   "2062_Warning_Data_BTCS_WARNING_WORD_13" : Word = PLC "2062_Warning_Data".BTCS_WARNING_WORD_13 AT %DB2062.DBW364, 1 s
   "2062_Warning_Data_BTCS_WARNING_WORD_14" : Word = PLC "2062_Warning_Data".BTCS_WARNING_WORD_14 AT %DB2062.DBW366, 1 s
   "2062_Warning_Data_BTCS_WARNING_WORD_15" : Word = PLC "2062_Warning_Data".BTCS_WARNING_WORD_15 AT %DB2062.DBW368, 1 s
   "2062_Warning_Data_BTCS_WARNING_WORD_16" : Word = PLC "2062_Warning_Data".BTCS_WARNING_WORD_16 AT %DB2062.DBW370, 1 s
   "2062_Warning_Data_BTCS_WARNING_WORD_2" : Word = PLC "2062_Warning_Data".BTCS_WARNING_WORD_02 AT %DB2062.DBW2, 1 s
   "2062_Warning_Data_BTCS_WARNING_WORD_3" : Word = PLC "2062_Warning_Data".BTCS_WARNING_WORD_03 AT %DB2062.DBW4, 1 s
   "2062_Warning_Data_BTCS_WARNING_WORD_4" : Word = PLC "2062_Warning_Data".BTCS_WARNING_WORD_04 AT %DB2062.DBW6, 1 s
   "2062_Warning_Data_BTCS_WARNING_WORD_5" : Word = PLC "2062_Warning_Data".BTCS_WARNING_WORD_05 AT %DB2062.DBW8, 1 s
   "2062_Warning_Data_BTCS_WARNING_WORD_6" : Word = PLC "2062_Warning_Data".BTCS_WARNING_WORD_06 AT %DB2062.DBW10, 1 s
   "2062_Warning_Data_BTCS_WARNING_WORD_7" : Word = PLC "2062_Warning_Data".BTCS_WARNING_WORD_07 AT %DB2062.DBW12, 1 s
   "2062_Warning_Data_BTCS_WARNING_WORD_8" : Word = PLC "2062_Warning_Data".BTCS_WARNING_WORD_08 AT %DB2062.DBW14, 1 s
   "2062_Warning_Data_Water Level Override 1P" : Bool = PLC "2062_Warning_Data"."Water Level Override 1P" AT %DB2062.DBX360.1, 1 s
   "2062_Warning_Data_Water Level Override 1S" : Bool = PLC "2062_Warning_Data"."Water Level Override 1S" AT %DB2062.DBX360.2, 1 s
   "2062_Warning_Data_Water Level Override 2P" : Bool = PLC "2062_Warning_Data"."Water Level Override 2P" AT %DB2062.DBX360.3, 1 s
   "2062_Warning_Data_Water Level Override 2S" : Bool = PLC "2062_Warning_Data"."Water Level Override 2S" AT %DB2062.DBX360.4, 1 s
   "2062_Warning_Data_Water Level Override 3P" : Bool = PLC "2062_Warning_Data"."Water Level Override 3P" AT %DB2062.DBX360.5, 1 s
   "2062_Warning_Data_Water Level Override 3S" : Bool = PLC "2062_Warning_Data"."Water Level Override 3S" AT %DB2062.DBX360.6, 1 s
   "2062_Warning_Data_Water Level Override 4P" : Bool = PLC "2062_Warning_Data"."Water Level Override 4P" AT %DB2062.DBX360.7, 1 s
   "2062_Warning_Data_Water Level Override 4S" : Bool = PLC "2062_Warning_Data"."Water Level Override 4S" AT %DB2062.DBX361.0, 1 s
   "2062_Warning_Data_Water Level Override 5P" : Bool = PLC "2062_Warning_Data"."Water Level Override 5P" AT %DB2062.DBX361.1, 1 s
   "2062_Warning_Data_Water Level Override 5S" : Bool = PLC "2062_Warning_Data"."Water Level Override 5S" AT %DB2062.DBX361.2, 1 s
   "2062_Warning_Data_Water Level Override 6P" : Bool = PLC "2062_Warning_Data"."Water Level Override 6P" AT %DB2062.DBX361.3, 1 s
   "2062_Warning_Data_Water Level Override 6S" : Bool = PLC "2062_Warning_Data"."Water Level Override 6S" AT %DB2062.DBX361.4, 1 s
   "2062_Warning_Data_Water Level Override APT" : Bool = PLC "2062_Warning_Data"."Water Level Override APT" AT %DB2062.DBX361.5, 1 s
   "2062_Warning_Data_Water Level Override FPT" : Bool = PLC "2062_Warning_Data"."Water Level Override FPT" AT %DB2062.DBX360.0, 1 s
   "2068_Sys_Status_Data_SAL_CNF_CHK" : Bool = PLC "2068_Sys_Status_Data".SAL_CNF_CHK, 100 ms
   "2068_Sys_Status_Data_SAL_VALID" : Bool = PLC "2068_Sys_Status_Data".SAL_VALID, 1 s
   "2086_Times_Alarm Enable Delay" : Time = PLC "2086_Times"."Alarm Enable Delay", 1 s
   "2086_Times_AT_DEOX_CNF_TIME" : Time = PLC "2086_Times".AT_DEOX_CNF_TIME AT %DB1.DBW0, 1 s
   "2086_Times_AT_REOX_CNF_TIME" : Time = PLC "2086_Times".AT_REOX_CNF_TIME AT %DB1.DBW0, 1 s
   "2086_Times_CV421_1S_MAX_TRVL_TIME" : Time = PLC "2086_Times".CV421_1S_MAX_TRVL_TIME, 1 s
   "2086_Times_CV421_2S_MAX_TRVL_TIME" : Time = PLC "2086_Times".CV421_2S_MAX_TRVL_TIME, 1 s
   "2086_Times_CV421_3S_MAX_TRVL_TIME" : Time = PLC "2086_Times".CV421_3S_MAX_TRVL_TIME, 1 s
   "2086_Times_CV421_4S_MAX_TRVL_TIME" : Time = PLC "2086_Times".CV421_4S_MAX_TRVL_TIME, 1 s
   "2086_Times_CV421_5S_MAX_TRVL_TIME" : Time = PLC "2086_Times".CV421_5S_MAX_TRVL_TIME, 1 s
   "2086_Times_CV421_6S_MAX_TRVL_TIME" : Time = PLC "2086_Times".CV421_6S_MAX_TRVL_TIME, 1 s
   "2086_Times_CV422_1P_MAX_TRVL_TIME" : Time = PLC "2086_Times".CV422_1P_MAX_TRVL_TIME, 1 s
   "2086_Times_CV422_2P_MAX_TRVL_TIME" : Time = PLC "2086_Times".CV422_2P_MAX_TRVL_TIME, 1 s
   "2086_Times_CV422_3P_MAX_TRVL_TIME" : Time = PLC "2086_Times".CV422_3P_MAX_TRVL_TIME, 1 s
   "2086_Times_CV422_4P_MAX_TRVL_TIME" : Time = PLC "2086_Times".CV422_4P_MAX_TRVL_TIME, 1 s
   "2086_Times_CV422_5P_MAX_TRVL_TIME" : Time = PLC "2086_Times".CV422_5P_MAX_TRVL_TIME, 1 s
   "2086_Times_CV422_6P_MAX_TRVL_TIME" : Time = PLC "2086_Times".CV422_6P_MAX_TRVL_TIME, 1 s
   "2086_Times_CV422_APT_MAX_TRVL_TIME" : Time = PLC "2086_Times".CV422_APT_MAX_TRVL_TIME, 1 s
   "2086_Times_CV422_FPT_MAX_TRVL_TIME" : Time = PLC "2086_Times".CV422_FPT_MAX_TRVL_TIME, 1 s
   "2086_Times_DEOX_PRE_GTT_CLS_DLY" : Time = PLC "2086_Times".DEOX_PRE_GTT_CLS_DLY AT %DB1.DBW0, 1 s
   "2086_Times_DEOX_PRE_GTT_OPN_DLY" : Time = PLC "2086_Times".DEOX_PRE_GTT_OPN_DLY AT %DB1.DBW0, 1 s
   "2086_Times_FIT417STAR Alarm Delay" : Time = PLC "2086_Times"."FIT417STAR Alarm Delay", 1 s
   "2086_Times_FIT418PORT Alarm Delay" : Time = PLC "2086_Times"."FIT418PORT Alarm Delay", 1 s
   "2086_Times_FIT419STAR Alarm Delay" : Time = PLC "2086_Times"."FIT419STAR Alarm Delay", 1 s
   "2086_Times_FIT420PORT Alarm Delay" : Time = PLC "2086_Times"."FIT420PORT Alarm Delay", 1 s
   "2086_Times_LS425 Port Alarm Delay" : Time = PLC "2086_Times"."LS425 Port Alarm Delay", 1 s
   "2086_Times_LS425 Star Alarm Delay" : Time = PLC "2086_Times"."LS425 Star Alarm Delay", 1 s
   "2086_Times_PIT424PORT Alarm Delay" : Time = PLC "2086_Times"."PIT424 Alarm Delay", 1 s
   "2086_Times_PS436 Alarm Delay" : Time = PLC "2086_Times"."PS436 Alarm Delay", 1 s
   "2086_Times_PT415PORT Alarm Delay" : Time = PLC "2086_Times"."PT415 Alarm Delay", 1 s
   "2086_Times_REOX_PRE_GTT_CLS_DLY" : Time = PLC "2086_Times".REOX_PRE_GTT_CLS_DLY AT %DB1.DBW0, 1 s
   "2086_Times_REOX_PRE_GTT_OPN_DLY" : Time = PLC "2086_Times".REOX_PRE_GTT_OPN_DLY AT %DB1.DBW0, 1 s
   "2086_Times_Tank Alarm Debounce" : Time = PLC "2086_Times"."Tank Alarm Reset Time", 1 s
   "2086_Times_TT426PORT Alarm Delay" : Time = PLC "2086_Times"."TT426_PORT_Alarm Delay", 1 s
   "2086_Times_TT426STAR Alarm Delay" : Time = PLC "2086_Times"."TT426_STAR_Alarm Delay", 1 s
   "21_FLOW_PRESSURE_SETPOINT_FIT_419_PRESSURE_SETPOINT" : Real = PLC "21_FLOW_PRESSURE_SETPOINT".FIT_419_PRESSURE_SETPOINT, 1 s
   "21_FLOW_PRESSURE_SETPOINT_FIT_420_PRESSURE_SETPOINT" : Real = PLC "21_FLOW_PRESSURE_SETPOINT".FIT_420_PRESSURE_SETPOINT, 1 s
   "2100_AUTO_SEQ_DB_SEQ_RNG" : Bool = PLC "2100_AUTO_SEQ_DB".SEQ_RNG, 1 s
   "2100_BTCS_CNTRL_DB_BTCS_STATE" : Int = PLC "2110_BTCS_CNTRL_DB".BTCS_STATE, 1 s
   "2100_BTCS_CNTRL_DB_BTCS_STEP" : Int = PLC "2110_BTCS_CNTRL_DB".BTCS_STEP, 1 s
   "2100_BTCS_CNTRL_DB_DE_OX_HRS" : Int = PLC "2110_BTCS_CNTRL_DB".DE_OX_HRS, 1 s
   "2100_BTCS_CNTRL_DB_DE_OX_MINS" : Int = PLC "2110_BTCS_CNTRL_DB".DE_OX_MINS, 1 s
   "2100_BTCS_CNTRL_DB_DE_OX_SP_HRS" : Int = PLC "2110_BTCS_CNTRL_DB".DE_OX_SP_HRS, 1 s
   "2100_BTCS_CNTRL_DB_DE_OX_SP_MINS" : Int = PLC "2110_BTCS_CNTRL_DB".DE_OX_SP_MINS, 1 s
   "2100_BTCS_CNTRL_DB_DWELL_HRS" : Int = PLC "2110_BTCS_CNTRL_DB".DWELL_HRS, 1 s
   "2100_BTCS_CNTRL_DB_DWELL_MINS" : Int = PLC "2110_BTCS_CNTRL_DB".DWELL_MINS, 1 s
   "2100_BTCS_CNTRL_DB_POST_DWELL_HRS" : Int = PLC "2110_BTCS_CNTRL_DB".POST_DWELL_HRS, 1 s
   "2100_BTCS_CNTRL_DB_POST_DWELL_MINS" : Int = PLC "2110_BTCS_CNTRL_DB".POST_DWELL_MINS, 1 s
   "2100_BTCS_CNTRL_DB_PRE_DWELL_HRS" : Int = PLC "2110_BTCS_CNTRL_DB".PRE_DWELL_HRS, 1 s
   "2100_BTCS_CNTRL_DB_PRE_DWELL_MINS" : Int = PLC "2110_BTCS_CNTRL_DB".PRE_DWELL_MINS, 1 s
   "2100_BTCS_CNTRL_DB_RE_OX_HRS" : Int = PLC "2110_BTCS_CNTRL_DB".RE_OX_HRS, 1 s
   "2100_BTCS_CNTRL_DB_RE_OX_MINS" : Int = PLC "2110_BTCS_CNTRL_DB".RE_OX_MINS, 1 s
   "2100_BTCS_CNTRL_DB_RE_OX_SP_HRS" : Int = PLC "2110_BTCS_CNTRL_DB".RE_OX_SP_HRS, 1 s
   "2100_BTCS_CNTRL_DB_RE_OX_SP_MINS" : Int = PLC "2110_BTCS_CNTRL_DB".RE_OX_SP_MINS, 1 s
   "2100_BTCS_CNTRL_DB_RMNG_SEQ_HRS" : Int = PLC "2110_BTCS_CNTRL_DB".RMNG_SEQ_HRS, 1 s
   "2100_BTCS_CNTRL_DB_RMNG_SEQ_MINS" : Int = PLC "2110_BTCS_CNTRL_DB".RMNG_SEQ_MINS, 1 s
   "2100_BTCS_CNTRL_DB_START_SEQ" : Bool = PLC "2110_BTCS_CNTRL_DB".START_SEQ, 1 s
   "2100_BTCS_CNTRL_DB_STOP_SEQ" : Bool = PLC "2110_BTCS_CNTRL_DB".STOP_SEQ, 1 s
   "2100_BTCS_CNTRL_DB_TOT_SEQ_HRS" : Int = PLC "2110_BTCS_CNTRL_DB".TOT_SEQ_HRS, 1 s
   "2100_BTCS_CNTRL_DB_TOT_SEQ_MINS" : Int = PLC "2110_BTCS_CNTRL_DB".TOT_SEQ_MINS, 1 s
   "2102_TIME_CALCS_DB_60X boost" : Bool = PLC "2102_TIME_CALCS_DB"."60X boost", 1 s
   "2102_TIME_CALCS_DB_DE_OX_MINS_RMNG" : Int = PLC "2102_TIME_CALCS_DB".DE_OX_MINS_RMNG, 1 s
   "2102_TIME_CALCS_DB_DE_OX_SP_MINS_RMNG" : Int = PLC "2102_TIME_CALCS_DB".DE_OX_SP_MINS_RMNG, 1 s
   "2102_TIME_CALCS_DB_DE_OX_SP_TMR_DN" : Bool = PLC "2102_TIME_CALCS_DB".DE_OX_SP_TMR_DN, 1 s
   "2102_TIME_CALCS_DB_DE_OX_TMR_DN" : Bool = PLC "2102_TIME_CALCS_DB".DE_OX_TMR_DN, 1 s
   "2102_TIME_CALCS_DB_DWELL_MINS_RMNG" : Int = PLC "2102_TIME_CALCS_DB".DWELL_MINS_RMNG, 1 s
   "2102_TIME_CALCS_DB_DWELL_TMR_DN" : Bool = PLC "2102_TIME_CALCS_DB".DWELL_TMR_DN, 1 s
   "2102_TIME_CALCS_DB_PHASE_DIFFERECE_MNS_REMNG" : Int = PLC "2102_TIME_CALCS_DB".PHASE_DIFFERECE_MNS_REMNG_De-Ox, 1 s
   "2102_TIME_CALCS_DB_POST_DWELL_MINS_RMNG" : Int = PLC "2102_TIME_CALCS_DB".POST_DWELL_MINS_RMNG, 1 s
   "2102_TIME_CALCS_DB_POST_DWELL_TMR_DN" : Bool = PLC "2102_TIME_CALCS_DB".POST_DWELL_TMR_DN, 1 s
   "2102_TIME_CALCS_DB_PRE_DWELL_MINS_RMNG" : Int = PLC "2102_TIME_CALCS_DB".PRE_DWELL_MINS_RMNG, 1 s
   "2102_TIME_CALCS_DB_PRE_DWELL_TMR_DN" : Bool = PLC "2102_TIME_CALCS_DB".PRE_DWELL_TMR_DN, 1 s
   "2102_TIME_CALCS_DB_PRE-DWEL MINS REMNG" : Int = PLC "2102_TIME_CALCS_DB"."PRE-DWEL MINS REMNG", 1 s
   "2102_TIME_CALCS_DB_PRE-DWEL_Warning 1" : Bool = PLC "2102_TIME_CALCS_DB"."PRE-DWEL_Warning 1", 500 ms
      on ChangeValue: "TimeRemainingToTreatment"()
   "2102_TIME_CALCS_DB_PRE-DWEL_Warning 2" : Bool = PLC "2102_TIME_CALCS_DB"."PRE-DWEL_Warning 2", 500 ms
      on ChangeValue: "TreatmentRequired"()
   "2102_TIME_CALCS_DB_PRE-DWEL_Warning 3" : Bool = PLC "2102_TIME_CALCS_DB"."PRE-DWEL_Warning 3", 1 s
   "2102_TIME_CALCS_DB_PRE-DWEL_Warning Min 1" : Int = PLC "2102_TIME_CALCS_DB"."PRE-DWEL_Warning Min 1", 1 s
   "2102_TIME_CALCS_DB_PRE-DWEL_Warning Min 2" : Int = PLC "2102_TIME_CALCS_DB"."PRE-DWEL_Warning Min 2", 1 s
   "2102_TIME_CALCS_DB_PRE-DWEL_Warning Min 3" : Int = PLC "2102_TIME_CALCS_DB"."PRE-DWEL_Warning Min 3", 1 s
   "2102_TIME_CALCS_DB_PRE-DWEL_Warning Reset 1" : Bool = PLC "2102_TIME_CALCS_DB"."PRE-DWEL_Warning Reset 1", 1 s
   "2102_TIME_CALCS_DB_PRE-DWEL_Warning Reset 2" : Bool = PLC "2102_TIME_CALCS_DB"."PRE-DWEL_Warning Reset 2", 1 s
   "2102_TIME_CALCS_DB_PRE-DWEL_Warning Reset 3" : Bool = PLC "2102_TIME_CALCS_DB"."PRE-DWEL_Warning Reset 3", 1 s
   "2102_TIME_CALCS_DB_RE_OX_MINS_RMNG" : Int = PLC "2102_TIME_CALCS_DB".RE_OX_MINS_RMNG, 1 s
   "2102_TIME_CALCS_DB_RE_OX_SP_MINS_RMNG" : Int = PLC "2102_TIME_CALCS_DB".RE_OX_SP_MINS_RMNG, 1 s
   "2102_TIME_CALCS_DB_RE_OX_SP_TMR_DN" : Bool = PLC "2102_TIME_CALCS_DB".RE_OX_SP_TMR_DN, 1 s
   "2102_TIME_CALCS_DB_RE_OX_TMR_DN" : Bool = PLC "2102_TIME_CALCS_DB".RE_OX_TMR_DN, 1 s
   "2102_TIME_CALCS_DB_Time_To_Treatment" : Int = PLC "2102_TIME_CALCS_DB".Time_To_Treatment, 1 s
   "2102_TIME_CALCS_DB_TIMES_VALID" : Bool = PLC "2102_TIME_CALCS_DB".TIMES_VALID, 1 s
   "2102_TIME_CALCS_DB_TOT_SEQ_DAYS" : Real = PLC "2102_TIME_CALCS_DB".TOT_SEQ_DAYS, 1 s
   "2102_TIME_CALCS_DB_TOT_SEQ_HRS_RMNG" : Int = PLC "2102_TIME_CALCS_DB".TOT_SEQ_HRS_RMNG, 1 s
   "2102_TIME_CALCS_DB_TOT_SEQ_MINS_RMNG" : Int = PLC "2102_TIME_CALCS_DB".TOT_SEQ_MINS_RMNG, 1 s
   "2102_TIME_CALCS_DB_Voyage_TIME_days" : Int = PLC "2102_TIME_CALCS_DB".Voyage_TIME_days, 1 s
   "2102_TIME_CALCS_DB_Voyage_TIME_hours" : Int = PLC "2102_TIME_CALCS_DB".Voyage_TIME_hours, 1 s
   "2102_TIME_CALCS_DB_Voyage_TIME_remaining_h" : Int = PLC "2102_TIME_CALCS_DB".Voyage_TIME_remaining_h, 1 s
   "2102_TIME_CALCS_DB_Voyage_TIME_remaining_m" : Int = PLC "2102_TIME_CALCS_DB".Voyage_TIME_remaining_m, 1 s
   "2110_BTCS_CNTRL_DB_PORT_TANK_STS" : Bool = PLC "2110_BTCS_CNTRL_DB".PORT_TANK_STS, 1 s
   "2110_BTCS_CNTRL_DB_RESET_ALL" : Bool = PLC "2110_BTCS_CNTRL_DB".RESET_ALL, 1 s
   "2110_BTCS_CNTRL_DB_STBD_TANK_STS" : Bool = PLC "2110_BTCS_CNTRL_DB".STBD_TANK_STS, 1 s
   "2115_VOYAGE_TIME_DAYS_VOYAGE_DAYS" : Real = PLC "2115_VOYAGE_TIME_DAYS".VOYAGE_DAYS, 1 s
   "40_TANKS_OP_DATA_RIO_02_VENT_A_2P" : Bool = PLC "40_TANKS_OP_DATA".RIO_02_VENT_A_2P AT %DB1.DBW0, 1 s
   "40_TANKS_OP_DATA_RIO_02_VENT_A_2S" : Bool = PLC "40_TANKS_OP_DATA".RIO_02_VENT_B_2S AT %DB1.DBW0, 1 s
   "40_TANKS_OP_DATA_RIO_02_VENT_B_2P" : Bool = PLC "40_TANKS_OP_DATA".RIO_02_VENT_B_2P AT %DB1.DBW0, 1 s
   "40_TANKS_OP_DATA_RIO_02_VENT_B_2S" : Bool = PLC "40_TANKS_OP_DATA".RIO_02_VENT_B_2P AT %DB1.DBW0, 1 s
   "502_ALM_ANALOG_IDB PIT 416_HIGH LEVEL VALUE (H)" : Real = PLC "502_ALM_ANALOG_IDB PIT 416"."HIGH LEVEL VALUE (H)" AT %DB65.DBD30, 1 s
   "502_ALM_ANALOG_IDB PIT 416_LOW LEVEL VALUE (L)" : Real = PLC "502_ALM_ANALOG_IDB PIT 416"."LOW LEVEL VALUE (L)" AT %DB65.DBD26, 1 s
   "502_ALM_ANALOG_IDB PIT 416_VERY HIGH LEVEL VALUE (HH)" : Real = PLC "502_ALM_ANALOG_IDB PIT 416"."VERY HIGH LEVEL VALUE (HH)" AT %DB65.DBD34, 1 s
   "502_ALM_ANALOG_IDB PIT 416_VERY LOW LEVEL VALUE (LL)" : Real = PLC "502_ALM_ANALOG_IDB PIT 416"."VERY LOW LEVEL VALUE (LL)" AT %DB65.DBD22, 1 s
   "503_WARNING CHCK_DB_2063_Alarm Word 12" : Word = PLC "503_WARNING CHCK_DB_2063"."Alarm Word 12", 1 s
   "503_WARNING CHCK_DB_2063_Alarm Word 13" : Word = PLC "503_WARNING CHCK_DB_2063"."Alarm Word 13", 1 s
   "503_WARNING CHCK_DB_2063_Alarm Word 14" : Word = PLC "503_WARNING CHCK_DB_2063"."Alarm Word 14", 1 s
   "503_WARNING CHCK_DB_2063_Alarm Word 15" : Word = PLC "503_WARNING CHCK_DB_2063"."Alarm Word 15", 1 s
   "503_WARNING CHCK_DB_2063_Alarm Word 16" : Word = PLC "503_WARNING CHCK_DB_2063"."Alarm Word 16", 1 s
   "504_Tank Grouping_DB2020_Boost" : Bool = PLC "504_Tank Grouping_DB2020".Boost, 1 s
   "504_Tank Grouping_DB2020_Cycle Length_ET" : Time = PLC "504_Tank Grouping_DB2020"."Cycle Length".ET, 1 s
   "504_Tank Grouping_DB2020_Cycle Period_ET" : Time = PLC "504_Tank Grouping_DB2020"."Cycle Period".ET, 1 s
   "504_Tank Grouping_DB2020_Diff Time Remain" : DInt = PLC "504_Tank Grouping_DB2020"."Diff Time Remain", 1 s
   "504_Tank Grouping_DB2020_GROUP ACTIV 1" : Bool = PLC "504_Tank Grouping_DB2020"."GROUP ACTIV 1", 1 s
   "504_Tank Grouping_DB2020_GROUP ACTIV 2" : Bool = PLC "504_Tank Grouping_DB2020"."GROUP ACTIV 2", 1 s
   "504_Tank Grouping_DB2020_GROUP ACTIV 3" : Bool = PLC "504_Tank Grouping_DB2020"."GROUP ACTIV 3", 1 s
   "504_Tank Grouping_DB2020_GROUP ACTIV 4" : Bool = PLC "504_Tank Grouping_DB2020"."GROUP ACTIV 4", 1 s
   "504_Tank Grouping_DB2020_GROUP ACTIV 5" : Bool = PLC "504_Tank Grouping_DB2020"."GROUP ACTIV 5", 1 s
   "504_Tank Grouping_DB2020_GROUP ACTIV 6" : Bool = PLC "504_Tank Grouping_DB2020"."GROUP ACTIV 6", 1 s
   "504_Tank Grouping_DB2020_GROUP ACTIV 7" : Bool = PLC "504_Tank Grouping_DB2020"."GROUP ACTIV 7", 1 s
   "504_Tank Grouping_DB2020_GROUP ACTIVE INT 1" : Bool = PLC "504_Tank Grouping_DB2020"."GROUP ACTIVE INT 1", 1 s
   "504_Tank Grouping_DB2020_GROUP ACTIVE INT 2" : Bool = PLC "504_Tank Grouping_DB2020"."GROUP ACTIVE INT 2", 1 s
   "504_Tank Grouping_DB2020_GROUP ACTIVE INT 3" : Bool = PLC "504_Tank Grouping_DB2020"."GROUP ACTIVE INT 3", 1 s
   "504_Tank Grouping_DB2020_GROUP ACTIVE INT 4" : Bool = PLC "504_Tank Grouping_DB2020"."GROUP ACTIVE INT 4", 1 s
   "504_Tank Grouping_DB2020_GROUP ACTIVE INT 5" : Bool = PLC "504_Tank Grouping_DB2020"."GROUP ACTIVE INT 5", 1 s
   "504_Tank Grouping_DB2020_GROUP ACTIVE INT 6" : Bool = PLC "504_Tank Grouping_DB2020"."GROUP ACTIVE INT 6", 1 s
   "504_Tank Grouping_DB2020_GROUP ACTIVE INT 7" : Bool = PLC "504_Tank Grouping_DB2020"."GROUP ACTIVE INT 7", 1 s
   "504_Tank Grouping_DB2020_GROUP of TANK 1" : Int = PLC "504_Tank Grouping_DB2020"."GROUP of TANK 1", 1 s
   "504_Tank Grouping_DB2020_GROUP of TANK 10" : Int = PLC "504_Tank Grouping_DB2020"."GROUP of TANK 10", 1 s
   "504_Tank Grouping_DB2020_GROUP of TANK 11" : Int = PLC "504_Tank Grouping_DB2020"."GROUP of TANK 11", 1 s
   "504_Tank Grouping_DB2020_GROUP of TANK 12" : Int = PLC "504_Tank Grouping_DB2020"."GROUP of TANK 12", 1 s
   "504_Tank Grouping_DB2020_GROUP of TANK 13" : Int = PLC "504_Tank Grouping_DB2020"."GROUP of TANK 13", 1 s
   "504_Tank Grouping_DB2020_GROUP of TANK 14" : Int = PLC "504_Tank Grouping_DB2020"."GROUP of TANK 14", 1 s
   "504_Tank Grouping_DB2020_GROUP of TANK 2" : Int = PLC "504_Tank Grouping_DB2020"."GROUP of TANK 2", 1 s
   "504_Tank Grouping_DB2020_GROUP of TANK 3" : Int = PLC "504_Tank Grouping_DB2020"."GROUP of TANK 3", 1 s
   "504_Tank Grouping_DB2020_GROUP of TANK 4" : Int = PLC "504_Tank Grouping_DB2020"."GROUP of TANK 4", 1 s
   "504_Tank Grouping_DB2020_GROUP of TANK 5" : Int = PLC "504_Tank Grouping_DB2020"."GROUP of TANK 5", 1 s
   "504_Tank Grouping_DB2020_GROUP of TANK 6" : Int = PLC "504_Tank Grouping_DB2020"."GROUP of TANK 6", 1 s
   "504_Tank Grouping_DB2020_GROUP of TANK 7" : Int = PLC "504_Tank Grouping_DB2020"."GROUP of TANK 7", 1 s
   "504_Tank Grouping_DB2020_GROUP of TANK 8" : Int = PLC "504_Tank Grouping_DB2020"."GROUP of TANK 8", 1 s
   "504_Tank Grouping_DB2020_GROUP of TANK 9" : Int = PLC "504_Tank Grouping_DB2020"."GROUP of TANK 9", 1 s
   "504_Tank Grouping_DB2020_GROUP SET" : Int = PLC "504_Tank Grouping_DB2020"."GROUP SET", 1 s
   "504_Tank Grouping_DB2020_O2 De-Ox Setpoint" : Real = PLC "504_Tank Grouping_DB2020"."O2 De-Ox Setpoint", 1 s
   "504_Tank Grouping_DB2020_Offset Timer_ET" : Time = PLC "504_Tank Grouping_DB2020"."Offset Timer".ET, 1 s
   "504_Tank Grouping_DB2020_RUN" : Bool = PLC "504_Tank Grouping_DB2020".RUN, 1 s
   "504_Tank Grouping_DB2020_RUN TANK 1" : Bool = PLC "504_Tank Grouping_DB2020"."RUN TANK 1", 1 s
   "504_Tank Grouping_DB2020_RUN TANK 10" : Bool = PLC "504_Tank Grouping_DB2020"."RUN TANK 10", 1 s
   "504_Tank Grouping_DB2020_RUN TANK 11" : Bool = PLC "504_Tank Grouping_DB2020"."RUN TANK 11", 1 s
   "504_Tank Grouping_DB2020_RUN TANK 12" : Bool = PLC "504_Tank Grouping_DB2020"."RUN TANK 12", 1 s
   "504_Tank Grouping_DB2020_RUN TANK 13" : Bool = PLC "504_Tank Grouping_DB2020"."RUN TANK 13", 1 s
   "504_Tank Grouping_DB2020_RUN TANK 14" : Bool = PLC "504_Tank Grouping_DB2020"."RUN TANK 14", 1 s
   "504_Tank Grouping_DB2020_RUN TANK 2" : Bool = PLC "504_Tank Grouping_DB2020"."RUN TANK 2", 1 s
   "504_Tank Grouping_DB2020_RUN TANK 3" : Bool = PLC "504_Tank Grouping_DB2020"."RUN TANK 3", 1 s
   "504_Tank Grouping_DB2020_RUN TANK 4" : Bool = PLC "504_Tank Grouping_DB2020"."RUN TANK 4", 1 s
   "504_Tank Grouping_DB2020_RUN TANK 5" : Bool = PLC "504_Tank Grouping_DB2020"."RUN TANK 5", 1 s
   "504_Tank Grouping_DB2020_RUN TANK 6" : Bool = PLC "504_Tank Grouping_DB2020"."RUN TANK 6", 1 s
   "504_Tank Grouping_DB2020_RUN TANK 7" : Bool = PLC "504_Tank Grouping_DB2020"."RUN TANK 7", 1 s
   "504_Tank Grouping_DB2020_RUN TANK 8" : Bool = PLC "504_Tank Grouping_DB2020"."RUN TANK 8", 1 s
   "504_Tank Grouping_DB2020_RUN TANK 9" : Bool = PLC "504_Tank Grouping_DB2020"."RUN TANK 9", 1 s
   "504_Tank Grouping_DB2020_Sequence Time Min Offset" : Time = PLC "504_Tank Grouping_DB2020"."Sequence Time m Offset", 1 s
   "504_Tank Grouping_DB2020_Sequence Time Min Offset_Int" : Real = PLC "504_Tank Grouping_DB2020"."Sequence Time m Offset_real", 1 s
   "504_Tank Grouping_DB2020_SetGroup" : Bool = PLC "504_Tank Grouping_DB2020".SetGroup, 1 s
   "504_Tank Grouping_DB2020_SetGroupSR" : Bool = PLC "504_Tank Grouping_DB2020".SetGroupSR, 1 s
   "504_Tank Grouping_DB2020_Tank1 Min Time_ET" : Time = PLC "504_Tank Grouping_DB2020"."Tank1 Min Time".ET, 1 s
   "504_Tank Grouping_DB2020_Tank10 Min Time_ET" : Time = PLC "504_Tank Grouping_DB2020"."Tank10 Min Time".ET, 1 s
   "504_Tank Grouping_DB2020_Tank12 Min Time_ET" : Time = PLC "504_Tank Grouping_DB2020"."Tank12 Min Time".ET, 1 s
   "504_Tank Grouping_DB2020_Tank13 Min Time_ET" : Time = PLC "504_Tank Grouping_DB2020"."Tank13 Min Time".ET, 1 s
   "504_Tank Grouping_DB2020_Tank14 Min Time_ET" : Time = PLC "504_Tank Grouping_DB2020"."Tank14 Min Time".ET, 1 s
   "504_Tank Grouping_DB2020_Tank2 Min Time_ET" : Time = PLC "504_Tank Grouping_DB2020"."Tank2 Min Time".ET, 1 s
   "504_Tank Grouping_DB2020_Tank3 Min Time_ET" : Time = PLC "504_Tank Grouping_DB2020"."Tank3 Min Time".ET, 1 s
   "504_Tank Grouping_DB2020_Tank4 Min Time_ET" : Time = PLC "504_Tank Grouping_DB2020"."Tank4 Min Time".ET, 1 s
   "504_Tank Grouping_DB2020_Tank5 Min Time_ET" : Time = PLC "504_Tank Grouping_DB2020"."Tank5 Min Time".ET, 1 s
   "504_Tank Grouping_DB2020_Tank6 Min Time_ET" : Time = PLC "504_Tank Grouping_DB2020"."Tank6 Min Time".ET, 1 s
   "504_Tank Grouping_DB2020_Tank7 Min Time_ET" : Time = PLC "504_Tank Grouping_DB2020"."Tank7 Min Time".ET, 1 s
   "504_Tank Grouping_DB2020_Tank8 Min Time_ET" : Time = PLC "504_Tank Grouping_DB2020"."Tank8 Min Time".ET, 1 s
   "504_Tank Grouping_DB2020_Tank9 Min Time_ET" : Time = PLC "504_Tank Grouping_DB2020"."Tank9 Min Time".ET, 1 s
   "504_Tank Grouping_DB2020_Time Left Tank_Time Left Tank 1" : Real = PLC "504_Tank Grouping_DB2020"."Time Left Tank"."Time Left Tank 1", 1 s
   "504_Tank Grouping_DB2020_Time Left Tank_Time Left Tank 10" : Real = PLC "504_Tank Grouping_DB2020"."Time Left Tank"."Time Left Tank 10", 1 s
   "504_Tank Grouping_DB2020_Time Left Tank_Time Left Tank 11" : Real = PLC "504_Tank Grouping_DB2020"."Time Left Tank"."Time Left Tank 11", 1 s
   "504_Tank Grouping_DB2020_Time Left Tank_Time Left Tank 12" : Real = PLC "504_Tank Grouping_DB2020"."Time Left Tank"."Time Left Tank 12", 1 s
   "504_Tank Grouping_DB2020_Time Left Tank_Time Left Tank 13" : Real = PLC "504_Tank Grouping_DB2020"."Time Left Tank"."Time Left Tank 13", 1 s
   "504_Tank Grouping_DB2020_Time Left Tank_Time Left Tank 14" : Real = PLC "504_Tank Grouping_DB2020"."Time Left Tank"."Time Left Tank 14", 1 s
   "504_Tank Grouping_DB2020_Time Left Tank_Time Left Tank 2" : Real = PLC "504_Tank Grouping_DB2020"."Time Left Tank"."Time Left Tank 2", 1 s
   "504_Tank Grouping_DB2020_Time Left Tank_Time Left Tank 3" : Real = PLC "504_Tank Grouping_DB2020"."Time Left Tank"."Time Left Tank 3", 1 s
   "504_Tank Grouping_DB2020_Time Left Tank_Time Left Tank 4" : Real = PLC "504_Tank Grouping_DB2020"."Time Left Tank"."Time Left Tank 4", 1 s
   "504_Tank Grouping_DB2020_Time Left Tank_Time Left Tank 5" : Real = PLC "504_Tank Grouping_DB2020"."Time Left Tank"."Time Left Tank 5", 1 s
   "504_Tank Grouping_DB2020_Time Left Tank_Time Left Tank 6" : Real = PLC "504_Tank Grouping_DB2020"."Time Left Tank"."Time Left Tank 6", 1 s
   "504_Tank Grouping_DB2020_Time Left Tank_Time Left Tank 7" : Real = PLC "504_Tank Grouping_DB2020"."Time Left Tank"."Time Left Tank 7", 1 s
   "504_Tank Grouping_DB2020_Time Left Tank_Time Left Tank 8" : Real = PLC "504_Tank Grouping_DB2020"."Time Left Tank"."Time Left Tank 8", 1 s
   "504_Tank Grouping_DB2020_Time Left Tank_Time Left Tank 9" : Real = PLC "504_Tank Grouping_DB2020"."Time Left Tank"."Time Left Tank 9", 1 s
   "504_Tank Grouping_DB2020_Valve Cycle_Enable" : Bool = PLC "504_Tank Grouping_DB2020"."Valve Cycle".Enable, 1 s
   "504_Tank Grouping_DB2020_Valve Cycle_Length" : Time = PLC "504_Tank Grouping_DB2020"."Valve Cycle".Length, 1 s
   "504_Tank Grouping_DB2020_Valve Cycle_Period" : Time = PLC "504_Tank Grouping_DB2020"."Valve Cycle".Period, 1 s
   "51_SLAVE_STATUS_RUNNING" : Bool = PLC "51_SLAVE_STATUS".RUNNING AT %DB51.DBX4.2, 1 s
   "60_Alarm_Data_ALRM_PRSNT" : Bool = PLC "60_Alarm_Data".ALRM_PRSNT AT %DB60.DBX32.0, 1 s
      on ChangeValue: "ALARM_Present"()
   "60_Alarm_Data_BC_ALARM_WORD_01" : Word = PLC "60_Alarm_Data".BC_ALARM_WORD_01 AT %DB60.DBW0, 1 s
   "60_Alarm_Data_BC_ALARM_WORD_02" : Word = PLC "60_Alarm_Data".BC_ALARM_WORD_02 AT %DB60.DBW2, 1 s
   "60_Alarm_Data_BC_ALARM_WORD_03" : Word = PLC "60_Alarm_Data".BC_ALARM_WORD_03 AT %DB60.DBW4, 1 s
   "60_Alarm_Data_BC_ALARM_WORD_04" : Word = PLC "60_Alarm_Data".BC_ALARM_WORD_04 AT %DB60.DBW6, 1 s
   "60_Alarm_Data_GCU_ALARM_WORD_01" : Word = PLC "60_Alarm_Data".GCU_ALARM_WORD_01 AT %DB60.DBW0, 1 s
   "60_Alarm_Data_GCU_ALARM_WORD_02" : Word = PLC "60_Alarm_Data".GCU_ALARM_WORD_02 AT %DB60.DBW2, 1 s
   "60_Alarm_Data_GCU_ALARM_WORD_03" : Word = PLC "60_Alarm_Data".GCU_ALARM_WORD_03 AT %DB60.DBW4, 1 s
   "60_Alarm_Data_GCU_ALARM_WORD_04" : Word = PLC "60_Alarm_Data".GCU_ALARM_WORD_04 AT %DB60.DBW6, 1 s
   "60_Alarm_Data_GCU_ALARM_WORD_05" : Word = PLC "60_Alarm_Data".GCU_ALARM_WORD_05 AT %DB60.DBW8, 1 s
   "60_Alarm_Data_GCU_ALARM_WORD_06" : Word = PLC "60_Alarm_Data".GCU_ALARM_WORD_06 AT %DB60.DBW10, 1 s
   "60_Alarm_Data_GCU_ALARM_WORD_07" : Word = PLC "60_Alarm_Data".GCU_ALARM_WORD_07 AT %DB60.DBW12, 1 s
   "60_Alarm_Data_GCU_ALARM_WORD_08" : Word = PLC "60_Alarm_Data".GCU_ALARM_WORD_08 AT %DB60.DBW14, 1 s
   "60_Alarm_Data_GCU_ALARM_WORD_09" : Word = PLC "60_Alarm_Data".GCU_ALARM_WORD_09 AT %DB60.DBW16, 1 s
   "60_Alarm_Data_IGG_ALARM_WORD_01" : Word = PLC "60_Alarm_Data".IGG_ALARM_WORD_01 AT %DB60.DBW0, 1 s
   "60_Alarm_Data_IGG_ALARM_WORD_02" : Word = PLC "60_Alarm_Data".IGG_ALARM_WORD_02 AT %DB60.DBW2, 1 s
   "60_Alarm_Data_IGG_ALARM_WORD_03" : Word = PLC "60_Alarm_Data".IGG_ALARM_WORD_03 AT %DB60.DBW4, 1 s
   "60_Alarm_Data_IGG_ALARM_WORD_04" : Word = PLC "60_Alarm_Data".IGG_ALARM_WORD_04 AT %DB60.DBW6, 1 s
   "62_Warning_Data_BC_WARNING_WORD_01" : Word = PLC "62_Warning_Data".BC_WARNING_WORD_01 AT %DB62.DBW0, 1 s
   "62_Warning_Data_BC_WARNING_WORD_02" : Word = PLC "62_Warning_Data".BC_WARNING_WORD_02 AT %DB62.DBW2, 1 s
   "62_Warning_Data_BC_WARNING_WORD_03" : Word = PLC "62_Warning_Data".BC_WARNING_WORD_03 AT %DB62.DBW4, 1 s
   "62_Warning_Data_BC_WARNING_WORD_04" : Word = PLC "62_Warning_Data".BC_WARNING_WORD_04 AT %DB62.DBW6, 1 s
   "62_Warning_Data_BC_WARNING_WORD_05" : Word = PLC "62_Warning_Data".BC_WARNING_WORD_05 AT %DB62.DBW8, 1 s
   "62_Warning_Data_BC_WARNING_WORD_06" : Word = PLC "62_Warning_Data".BC_WARNING_WORD_06 AT %DB62.DBW10, 1 s
   "62_Warning_Data_GCU_WARNING_WORD_01" : Word = PLC "62_Warning_Data".GCU_WARNING_WORD_01 AT %DB62.DBW0, 1 s
   "62_Warning_Data_GCU_WARNING_WORD_02" : Word = PLC "62_Warning_Data".GCU_WARNING_WORD_02 AT %DB62.DBW2, 1 s
   "62_Warning_Data_GCU_WARNING_WORD_03" : Word = PLC "62_Warning_Data".GCU_WARNING_WORD_03 AT %DB62.DBW4, 1 s
   "62_Warning_Data_GCU_WARNING_WORD_04" : Word = PLC "62_Warning_Data".GCU_WARNING_WORD_04 AT %DB62.DBW6, 1 s
   "62_Warning_Data_GCU_WARNING_WORD_05" : Word = PLC "62_Warning_Data".GCU_WARNING_WORD_05 AT %DB62.DBW8, 1 s
   "62_Warning_Data_GCU_WARNING_WORD_06" : Word = PLC "62_Warning_Data".GCU_WARNING_WORD_06 AT %DB62.DBW10, 1 s
   "62_Warning_Data_GCU_WARNING_WORD_07" : Word = PLC "62_Warning_Data".GCU_WARNING_WORD_07 AT %DB62.DBW12, 1 s
   "62_Warning_Data_GCU_WARNING_WORD_08" : Word = PLC "62_Warning_Data".GCU_WARNING_WORD_08 AT %DB62.DBW14, 1 s
   "62_Warning_Data_GCU_WARNING_WORD_09" : Word = PLC "62_Warning_Data".GCU_WARNING_WORD_09 AT %DB62.DBW16, 1 s
   "62_Warning_Data_IGG_WARNING_WORD_01" : Word = PLC "62_Warning_Data".IGG_WARNING_WORD_01 AT %DB62.DBW0, 1 s
   "62_Warning_Data_IGG_WARNING_WORD_02" : Word = PLC "62_Warning_Data".IGG_WARNING_WORD_02 AT %DB62.DBW2, 1 s
   "62_Warning_Data_IGG_WARNING_WORD_03" : Word = PLC "62_Warning_Data".IGG_WARNING_WORD_03 AT %DB62.DBW4, 1 s
   "62_Warning_Data_IGG_WARNING_WORD_04" : Word = PLC "62_Warning_Data".IGG_WARNING_WORD_04 AT %DB62.DBW6, 1 s
   "62_Warning_Data_IGG_WARNING_WORD_05" : Word = PLC "62_Warning_Data".IGG_WARNING_WORD_05 AT %DB62.DBW8, 1 s
   "62_Warning_Data_IGG_WARNING_WORD_06" : Word = PLC "62_Warning_Data".IGG_WARNING_WORD_06 AT %DB62.DBW10, 1 s
   "62_Warning_Data_WRNG_PRSNT" : Bool = PLC "62_Warning_Data".WRNG_PRSNT AT %DB62.DBX16.0, 1 s
   "64_Functioning Hours_E500A_IDB_Hours Functioning" : Int = PLC "64_Functioning Hours_E500A_IDB"."Hours Functioning", 1 s
   "64_Functioning Hours_E500B_IDB_Hours Functioning" : Int = PLC "64_Functioning Hours_E500B_IDB"."Hours Functioning", 1 s
   "64_Functioning Hours_P301_IDB_Hours Functioning" : Int = PLC "64_Functioning Hours_P301_IDB"."Hours Functioning", 1 s
   "64_Message_Data_BC_MESSAGE_WORD_01" : Word = PLC "64_Message_Data".BC_MESSAGE_WORD_01 AT %DB64.DBW0, 1 s
   "64_Message_Data_BC_MESSAGE_WORD_02" : Word = PLC "64_Message_Data".BC_MESSAGE_WORD_02 AT %DB64.DBW2, 1 s
   "64_Message_Data_IGG_MESSAGE_WORD_01" : Word = PLC "64_Message_Data".IGG_MESSAGE_WORD_01 AT %DB64.DBW0, 1 s
   "64_Message_Data_IGG_MESSAGE_WORD_02" : Word = PLC "64_Message_Data".IGG_MESSAGE_WORD_02 AT %DB64.DBW2, 1 s
   "66_Event_Data_BC_EVENT_WORD_01" : Word = PLC "66_Event_Data".BC_EVENT_WORD_01 AT %DB66.DBW0, 1 s
   "66_Event_Data_BC_EVENT_WORD_02" : Word = PLC "66_Event_Data".BC_EVENT_WORD_02 AT %DB66.DBW2, 1 s
   "66_Event_Data_IGG_EVENT_WORD_01" : Word = PLC "66_Event_Data".IGG_EVENT_WORD_01 AT %DB66.DBW0, 1 s
   "66_Event_Data_IGG_EVENT_WORD_02" : Word = PLC "66_Event_Data".IGG_EVENT_WORD_02 AT %DB66.DBW2, 1 s
   "68_Sys_Status_Data_FUEL_PRES_IN_RNG" : Bool = PLC "68_Sys_Status_Data".FUEL_PRES_IN_RNG, 1 s
   "68_Sys_Status_Data_IA_PRES_IN_RNG" : Bool = PLC "68_Sys_Status_Data".IA_PRES_IN_RNG, 1 s
   "68_Sys_Status_Data_INTRLKS_OK" : Bool = PLC "68_Sys_Status_Data".INTRLKS_OK, 1 s
   "70_Mode_Data_AUT_RST_PLS_IN" : Bool = PLC "70_Mode_Data".AUT_RST_PLS.IN, 1 s
   "7T1 Power Healthy" : Bool = PLC "10_DI_Data".7T1_PWR_OK AT %DB1.DBX0.0, 1 s
   "7T2 Power Healthy" : Bool = PLC "10_DI_Data".7T2_PWR_OK AT %DB1.DBX0.0, 1 s
   "7T3 Power Healthy" : Bool = PLC "10_DI_Data".7T3_PWR_OK AT %DB1.DBX0.0, 1 s
   "80_From_HMI_Beacon frequency" : Time = PLC "80_From_HMI"."Beacon frequency", 1 s
   "80_From_HMI_BurnerProgramedStop" : Bool = PLC "80_From_HMI".BurnerProgramedStop, 1 s
   "80_From_HMI_Buzzer reset time" : Time = PLC "80_From_HMI"."Buzzer reset time", 1 s
   "80_From_HMI_FLM_FAIL_DLY" : Time = PLC "80_From_HMI".FLM_FAIL_DLY, 1 s
   "80_From_HMI_FS317 delay" : Time = PLC "86_Times"."FS317 delay", 1 s
   "80_From_HMI_FS320 delay" : Time = PLC "86_Times"."FS320 delay", 1 s
   "80_From_HMI_FS332 Delay" : Time = PLC "86_Times"."FS332 Delay", 1 s
   "80_From_HMI_LOW_SAL_ACPT" : Bool = PLC "80_From_HMI".LOW_SAL_ACPT, 1 s
   "80_From_HMI_LOW_SAL_RJCT" : Bool = PLC "80_From_HMI".LOW_SAL_RJCT, 1 s
   "80_From_HMI_MAN_AQ_DEC_800" : Bool = PLC "80_From_HMI".MAN_AQ_DEC_800, 1 s
   "80_From_HMI_MAN_AQ_DEC_802" : Bool = PLC "80_From_HMI".MAN_AQ_DEC_802, 1 s
   "80_From_HMI_MAN_AQ_DEC_804" : Bool = PLC "80_From_HMI".MAN_AQ_DEC_804, 1 s
   "80_From_HMI_MAN_AQ_DEC_806" : Bool = PLC "80_From_HMI".MAN_AQ_DEC_806, 1 s
   "80_From_HMI_MAN_AQ_INC_800" : Bool = PLC "80_From_HMI".MAN_AQ_INC_800, 1 s
   "80_From_HMI_MAN_AQ_INC_802" : Bool = PLC "80_From_HMI".MAN_AQ_INC_802, 1 s
   "80_From_HMI_MAN_AQ_INC_804" : Bool = PLC "80_From_HMI".MAN_AQ_INC_804, 1 s
   "80_From_HMI_MAN_AQ_INC_806" : Bool = PLC "80_From_HMI".MAN_AQ_INC_806, 1 s
   "80_From_HMI_MAN_DQ_136_0" : Bool = PLC "80_From_HMI".MAN_DQ_136_0, 1 s
   "80_From_HMI_MAN_DQ_136_1" : Bool = PLC "80_From_HMI".MAN_DQ_136_1, 1 s
   "80_From_HMI_MAN_DQ_136_2" : Bool = PLC "80_From_HMI".MAN_DQ_136_2, 1 s
   "80_From_HMI_MAN_DQ_136_3" : Bool = PLC "80_From_HMI".MAN_DQ_136_3, 1 s
   "80_From_HMI_MAN_DQ_136_4" : Bool = PLC "80_From_HMI".MAN_DQ_136_4, 1 s
   "80_From_HMI_MAN_DQ_136_5" : Bool = PLC "80_From_HMI".MAN_DQ_136_5, 1 s
   "80_From_HMI_MAN_DQ_136_6" : Bool = PLC "80_From_HMI".MAN_DQ_136_6, 1 s
   "80_From_HMI_MAN_DQ_136_7" : Bool = PLC "80_From_HMI".MAN_DQ_136_7, 1 s
   "80_From_HMI_MAN_DQ_137_0" : Bool = PLC "80_From_HMI".MAN_DQ_137_0, 1 s
   "80_From_HMI_MAN_DQ_137_1" : Bool = PLC "80_From_HMI".MAN_DQ_137_1, 1 s
   "80_From_HMI_MAN_DQ_137_2" : Bool = PLC "80_From_HMI".MAN_DQ_137_2, 1 s
   "80_From_HMI_MAN_DQ_137_3" : Bool = PLC "80_From_HMI".MAN_DQ_137_3, 1 s
   "80_From_HMI_MAN_DQ_137_4" : Bool = PLC "80_From_HMI".MAN_DQ_137_4, 1 s
   "80_From_HMI_MAN_DQ_137_5" : Bool = PLC "80_From_HMI".MAN_DQ_137_5, 1 s
   "80_From_HMI_MAN_DQ_137_6" : Bool = PLC "80_From_HMI".MAN_DQ_137_6, 1 s
   "80_From_HMI_MAN_DQ_137_7" : Bool = PLC "80_From_HMI".MAN_DQ_137_7, 1 s
   "80_From_HMI_MAN_DQ_138_0" : Bool = PLC "80_From_HMI".MAN_DQ_138_0, 1 s
   "80_From_HMI_MAN_DQ_138_1" : Bool = PLC "80_From_HMI".MAN_DQ_138_1, 1 s
   "80_From_HMI_MAN_DQ_138_2" : Bool = PLC "80_From_HMI".MAN_DQ_138_2, 1 s
   "80_From_HMI_MAN_DQ_138_3" : Bool = PLC "80_From_HMI".MAN_DQ_138_3, 1 s
   "80_From_HMI_MAN_DQ_138_4" : Bool = PLC "80_From_HMI".MAN_DQ_138_4, 1 s
   "80_From_HMI_MAN_DQ_138_5" : Bool = PLC "80_From_HMI".MAN_DQ_138_5, 1 s
   "80_From_HMI_MAN_DQ_138_6" : Bool = PLC "80_From_HMI".MAN_DQ_138_6, 1 s
   "80_From_HMI_MAN_DQ_138_7" : Bool = PLC "80_From_HMI".MAN_DQ_138_7, 1 s
   "80_From_HMI_MAN_DQ_139_0" : Bool = PLC "80_From_HMI".MAN_DQ_139_0, 1 s
   "80_From_HMI_MAN_DQ_139_1" : Bool = PLC "80_From_HMI".MAN_DQ_139_1, 1 s
   "80_From_HMI_MAN_DQ_139_2" : Bool = PLC "80_From_HMI".MAN_DQ_139_2, 1 s
   "80_From_HMI_MAN_DQ_139_3" : Bool = PLC "80_From_HMI".MAN_DQ_139_3, 1 s